REGION Network 3
   RUNG wire#powerrail
      Move(in := "EMS".Carrier[#Carrier].Zone, out1 => #Zone_Echo)
   END_RUNG
   // the same network as SCL:
   #Zone_Echo := "EMS".Carrier[#Carrier].Zone;
END_REGION

REGION Network 4
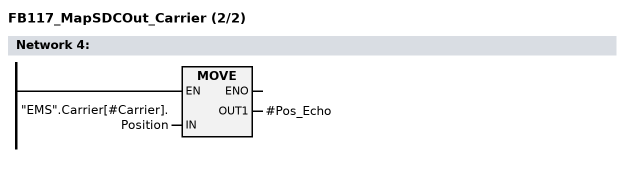
   RUNG wire#powerrail
      Move(in := "EMS".Carrier[#Carrier].Position, out1 => #Pos_Echo)
   END_RUNG
   // the same network as SCL:
   #Pos_Echo := "EMS".Carrier[#Carrier].Position;
END_REGION
END_FUNCTION_BLOCK

FUNCTION_BLOCK "FB118_TCMapSDCOut"   // FB118, LAD
{ S7_Optimized_Access := 'TRUE' }
VERSION : 0.1
   VAR_INPUT
      TC_ZoneMotion : "UDT_TC_ZoneMotion";
      Zone : Int;
      Carrier : Int;
   END_VAR
   VAR_OUTPUT
      SDCOUT_DriveFwdCmd : Bool;
      SDCOUT_DriveCmdSpeed : Word;
      SDCOUT_NextStopPos : DWord;
      SDCOUT_NextCarrierNum : Word;
      SDCOut_AtCmdPos : Bool;
   END_VAR
   VAR
      CarrierTempZone : Int;
      oneshot : Array[0..20] of Bool;
      oneshotneg : Bool;
      oneshot3 : Bool;
      resetlatch1 : Bool;
      DriveCmdSetup : Array[0..99] of Bool;
   END_VAR
   VAR_TEMP
      tempptrig : Bool;
   END_VAR
BEGIN

REGION Network 1
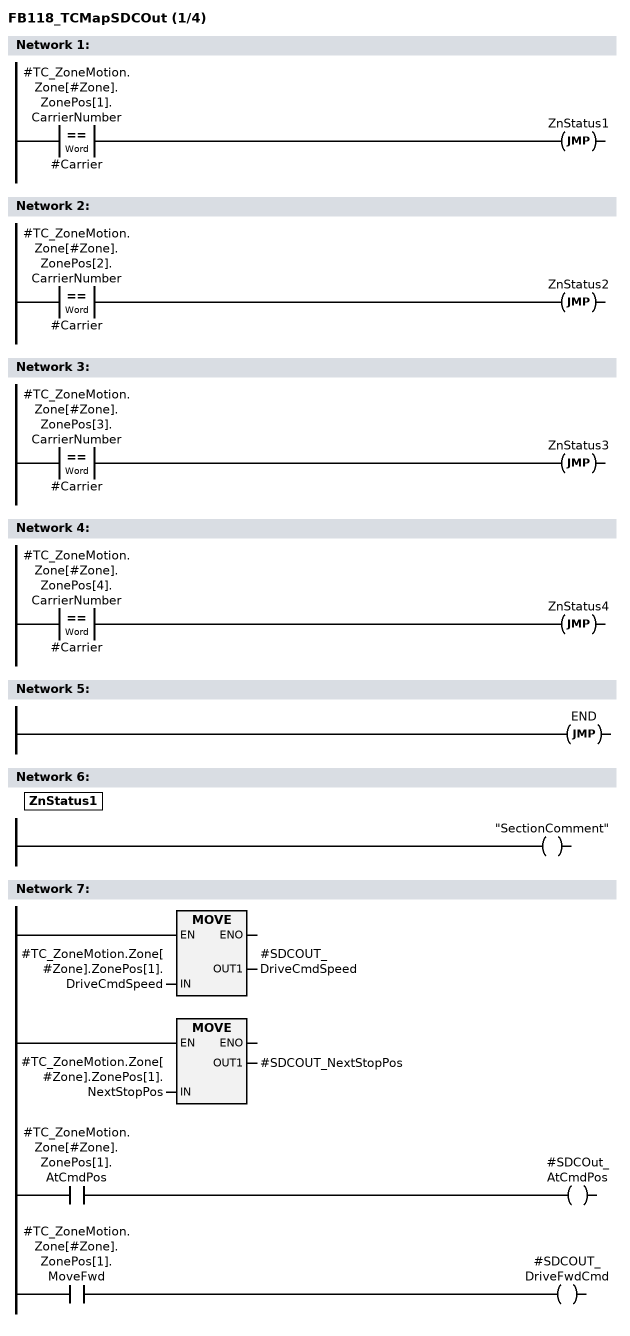
   RUNG wire#powerrail
      { S7_Templates := "SrcType := Word" } EQ_Contact(in1 := #TC_ZoneMotion.Zone[#Zone].ZonePos[1].CarrierNumber, in2 := #Carrier)
      JumpCoil( ZnStatus1 )
   END_RUNG
   // the same network as SCL:
   IF #TC_ZoneMotion.Zone[#Zone].ZonePos[1].CarrierNumber = #Carrier THEN GOTO ZnStatus1; END_IF;
END_REGION

REGION Network 2
   RUNG wire#powerrail
      { S7_Templates := "SrcType := Word" } EQ_Contact(in1 := #TC_ZoneMotion.Zone[#Zone].ZonePos[2].CarrierNumber, in2 := #Carrier)
      JumpCoil( ZnStatus2 )
   END_RUNG
   // the same network as SCL:
   IF #TC_ZoneMotion.Zone[#Zone].ZonePos[2].CarrierNumber = #Carrier THEN GOTO ZnStatus2; END_IF;
END_REGION

REGION Network 3
   RUNG wire#powerrail
      { S7_Templates := "SrcType := Word" } EQ_Contact(in1 := #TC_ZoneMotion.Zone[#Zone].ZonePos[3].CarrierNumber, in2 := #Carrier)
      JumpCoil( ZnStatus3 )
   END_RUNG
   // the same network as SCL:
   IF #TC_ZoneMotion.Zone[#Zone].ZonePos[3].CarrierNumber = #Carrier THEN GOTO ZnStatus3; END_IF;
END_REGION

REGION Network 4
   RUNG wire#powerrail
      { S7_Templates := "SrcType := Word" } EQ_Contact(in1 := #TC_ZoneMotion.Zone[#Zone].ZonePos[4].CarrierNumber, in2 := #Carrier)
      JumpCoil( ZnStatus4 )
   END_RUNG
   // the same network as SCL:
   IF #TC_ZoneMotion.Zone[#Zone].ZonePos[4].CarrierNumber = #Carrier THEN GOTO ZnStatus4; END_IF;
END_REGION

REGION Network 5
   RUNG wire#powerrail
      JumpCoil( END )
   END_RUNG
   // the same network as SCL:
   GOTO END;
END_REGION

REGION Network 6
   Label( ZnStatus1 )
   RUNG wire#powerrail
      Coil( "SectionComment" )
   END_RUNG
   // the same network as SCL:
   ZnStatus1:
   "SectionComment" := TRUE;
END_REGION

REGION Network 7
   RUNG wire#powerrail
      Move(in := #TC_ZoneMotion.Zone[#Zone].ZonePos[1].DriveCmdSpeed, out1 => #SDCOUT_DriveCmdSpeed)
   END_RUNG
   RUNG wire#powerrail
      Move(in := #TC_ZoneMotion.Zone[#Zone].ZonePos[1].NextStopPos, out1 => #SDCOUT_NextStopPos)
   END_RUNG
   RUNG wire#powerrail
      Contact( #TC_ZoneMotion.Zone[#Zone].ZonePos[1].AtCmdPos )
      Coil( #SDCOut_AtCmdPos )
   END_RUNG
   RUNG wire#powerrail
      Contact( #TC_ZoneMotion.Zone[#Zone].ZonePos[1].MoveFwd )
      Coil( #SDCOUT_DriveFwdCmd )
   END_RUNG
   // the same network as SCL:
   #SDCOUT_DriveCmdSpeed := #TC_ZoneMotion.Zone[#Zone].ZonePos[1].DriveCmdSpeed;
   #SDCOUT_NextStopPos := #TC_ZoneMotion.Zone[#Zone].ZonePos[1].NextStopPos;
   #SDCOut_AtCmdPos := #TC_ZoneMotion.Zone[#Zone].ZonePos[1].AtCmdPos;
   #SDCOUT_DriveFwdCmd := #TC_ZoneMotion.Zone[#Zone].ZonePos[1].MoveFwd;
END_REGION

REGION Network 8
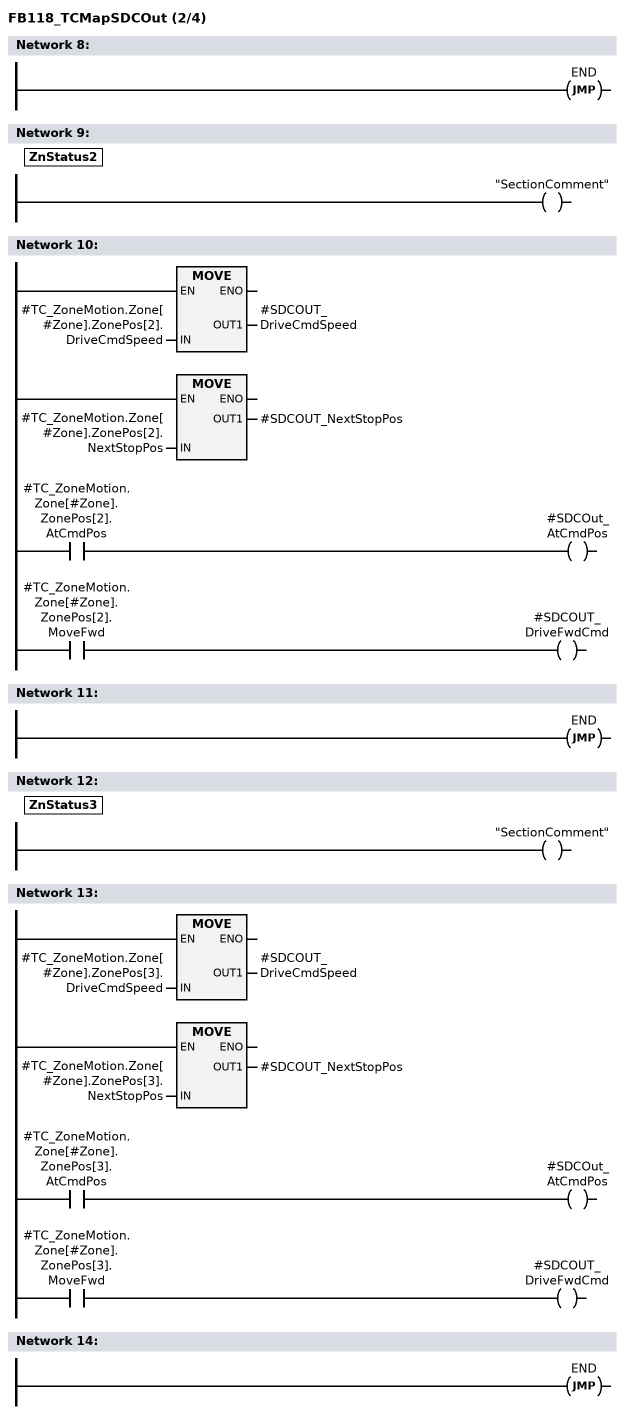
   RUNG wire#powerrail
      JumpCoil( END )
   END_RUNG
   // the same network as SCL:
   GOTO END;
END_REGION

REGION Network 9
   Label( ZnStatus2 )
   RUNG wire#powerrail
      Coil( "SectionComment" )
   END_RUNG
   // the same network as SCL:
   ZnStatus2:
   "SectionComment" := TRUE;
END_REGION

REGION Network 10
   RUNG wire#powerrail
      Move(in := #TC_ZoneMotion.Zone[#Zone].ZonePos[2].DriveCmdSpeed, out1 => #SDCOUT_DriveCmdSpeed)
   END_RUNG
   RUNG wire#powerrail
      Move(in := #TC_ZoneMotion.Zone[#Zone].ZonePos[2].NextStopPos, out1 => #SDCOUT_NextStopPos)
   END_RUNG
   RUNG wire#powerrail
      Contact( #TC_ZoneMotion.Zone[#Zone].ZonePos[2].AtCmdPos )
      Coil( #SDCOut_AtCmdPos )
   END_RUNG
   RUNG wire#powerrail
      Contact( #TC_ZoneMotion.Zone[#Zone].ZonePos[2].MoveFwd )
      Coil( #SDCOUT_DriveFwdCmd )
   END_RUNG
   // the same network as SCL:
   #SDCOUT_DriveCmdSpeed := #TC_ZoneMotion.Zone[#Zone].ZonePos[2].DriveCmdSpeed;
   #SDCOUT_NextStopPos := #TC_ZoneMotion.Zone[#Zone].ZonePos[2].NextStopPos;
   #SDCOut_AtCmdPos := #TC_ZoneMotion.Zone[#Zone].ZonePos[2].AtCmdPos;
   #SDCOUT_DriveFwdCmd := #TC_ZoneMotion.Zone[#Zone].ZonePos[2].MoveFwd;
END_REGION

REGION Network 11
   RUNG wire#powerrail
      JumpCoil( END )
   END_RUNG
   // the same network as SCL:
   GOTO END;
END_REGION

REGION Network 12
   Label( ZnStatus3 )
   RUNG wire#powerrail
      Coil( "SectionComment" )
   END_RUNG
   // the same network as SCL:
   ZnStatus3:
   "SectionComment" := TRUE;
END_REGION

REGION Network 13
   RUNG wire#powerrail
      Move(in := #TC_ZoneMotion.Zone[#Zone].ZonePos[3].DriveCmdSpeed, out1 => #SDCOUT_DriveCmdSpeed)
   END_RUNG
   RUNG wire#powerrail
      Move(in := #TC_ZoneMotion.Zone[#Zone].ZonePos[3].NextStopPos, out1 => #SDCOUT_NextStopPos)
   END_RUNG
   RUNG wire#powerrail
      Contact( #TC_ZoneMotion.Zone[#Zone].ZonePos[3].AtCmdPos )
      Coil( #SDCOut_AtCmdPos )
   END_RUNG
   RUNG wire#powerrail
      Contact( #TC_ZoneMotion.Zone[#Zone].ZonePos[3].MoveFwd )
      Coil( #SDCOUT_DriveFwdCmd )
   END_RUNG
   // the same network as SCL:
   #SDCOUT_DriveCmdSpeed := #TC_ZoneMotion.Zone[#Zone].ZonePos[3].DriveCmdSpeed;
   #SDCOUT_NextStopPos := #TC_ZoneMotion.Zone[#Zone].ZonePos[3].NextStopPos;
   #SDCOut_AtCmdPos := #TC_ZoneMotion.Zone[#Zone].ZonePos[3].AtCmdPos;
   #SDCOUT_DriveFwdCmd := #TC_ZoneMotion.Zone[#Zone].ZonePos[3].MoveFwd;
END_REGION

REGION Network 14
   RUNG wire#powerrail
      JumpCoil( END )
   END_RUNG
   // the same network as SCL:
   GOTO END;
END_REGION

REGION Network 15
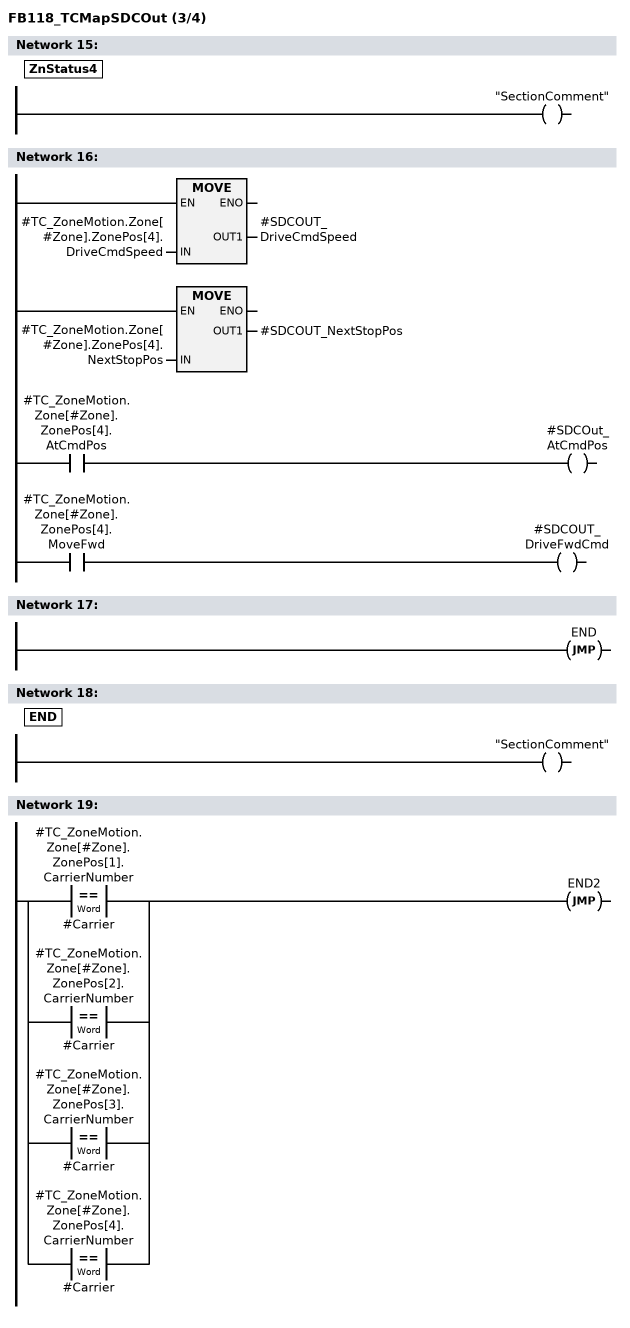
   Label( ZnStatus4 )
   RUNG wire#powerrail
      Coil( "SectionComment" )
   END_RUNG
   // the same network as SCL:
   ZnStatus4:
   "SectionComment" := TRUE;
END_REGION

REGION Network 16
   RUNG wire#powerrail
      Move(in := #TC_ZoneMotion.Zone[#Zone].ZonePos[4].DriveCmdSpeed, out1 => #SDCOUT_DriveCmdSpeed)
   END_RUNG
   RUNG wire#powerrail
      Move(in := #TC_ZoneMotion.Zone[#Zone].ZonePos[4].NextStopPos, out1 => #SDCOUT_NextStopPos)
   END_RUNG
   RUNG wire#powerrail
      Contact( #TC_ZoneMotion.Zone[#Zone].ZonePos[4].AtCmdPos )
      Coil( #SDCOut_AtCmdPos )
   END_RUNG
   RUNG wire#powerrail
      Contact( #TC_ZoneMotion.Zone[#Zone].ZonePos[4].MoveFwd )
      Coil( #SDCOUT_DriveFwdCmd )
   END_RUNG
   // the same network as SCL:
   #SDCOUT_DriveCmdSpeed := #TC_ZoneMotion.Zone[#Zone].ZonePos[4].DriveCmdSpeed;
   #SDCOUT_NextStopPos := #TC_ZoneMotion.Zone[#Zone].ZonePos[4].NextStopPos;
   #SDCOut_AtCmdPos := #TC_ZoneMotion.Zone[#Zone].ZonePos[4].AtCmdPos;
   #SDCOUT_DriveFwdCmd := #TC_ZoneMotion.Zone[#Zone].ZonePos[4].MoveFwd;
END_REGION

REGION Network 17
   RUNG wire#powerrail
      JumpCoil( END )
   END_RUNG
   // the same network as SCL:
   GOTO END;
END_REGION

REGION Network 18
   Label( END )
   RUNG wire#powerrail
      Coil( "SectionComment" )
   END_RUNG
   // the same network as SCL:
   END:
   "SectionComment" := TRUE;
END_REGION

REGION Network 19
   RUNG wire#powerrail
      { S7_Templates := "SrcType := Word" } EQ_Contact(in1 := #TC_ZoneMotion.Zone[#Zone].ZonePos[1].CarrierNumber, in2 := #Carrier)
      wire#w1
      JumpCoil( END2 )
   END_RUNG
   RUNG wire#powerrail
      { S7_Templates := "SrcType := Word" } EQ_Contact(in1 := #TC_ZoneMotion.Zone[#Zone].ZonePos[2].CarrierNumber, in2 := #Carrier)
   END_RUNG wire#w1
   RUNG wire#powerrail
      { S7_Templates := "SrcType := Word" } EQ_Contact(in1 := #TC_ZoneMotion.Zone[#Zone].ZonePos[3].CarrierNumber, in2 := #Carrier)
   END_RUNG wire#w1
   RUNG wire#powerrail
      { S7_Templates := "SrcType := Word" } EQ_Contact(in1 := #TC_ZoneMotion.Zone[#Zone].ZonePos[4].CarrierNumber, in2 := #Carrier)
   END_RUNG wire#w1
   // the same network as SCL:
   IF (#TC_ZoneMotion.Zone[#Zone].ZonePos[1].CarrierNumber = #Carrier) OR (#TC_ZoneMotion.Zone[#Zone].ZonePos[2].CarrierNumber = #Carrier) OR (#TC_ZoneMotion.Zone[#Zone].ZonePos[3].CarrierNumber = #Carrier) OR (#TC_ZoneMotion.Zone[#Zone].ZonePos[4].CarrierNumber = #Carrier) THEN
       GOTO END2;
   END_IF;
END_REGION

REGION Network 20
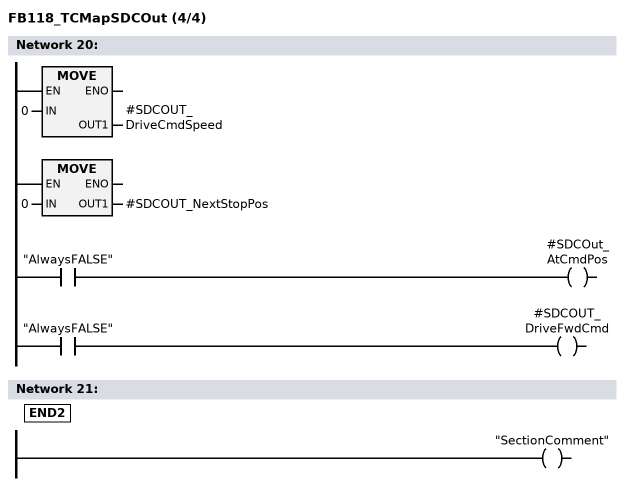
   RUNG wire#powerrail
      Move(in := 0, out1 => #SDCOUT_DriveCmdSpeed)
   END_RUNG
   RUNG wire#powerrail
      Move(in := 0, out1 => #SDCOUT_NextStopPos)
   END_RUNG
   RUNG wire#powerrail
      Contact( "AlwaysFALSE" )
      Coil( #SDCOut_AtCmdPos )
   END_RUNG
   RUNG wire#powerrail
      Contact( "AlwaysFALSE" )
      Coil( #SDCOUT_DriveFwdCmd )
   END_RUNG
   // the same network as SCL:
   #SDCOUT_DriveCmdSpeed := 0;
   #SDCOUT_NextStopPos := 0;
   #SDCOut_AtCmdPos := "AlwaysFALSE";
   #SDCOUT_DriveFwdCmd := "AlwaysFALSE";
END_REGION

REGION Network 21
   Label( END2 )
   RUNG wire#powerrail
      Coil( "SectionComment" )
   END_RUNG
   // the same network as SCL:
   END2:
   "SectionComment" := TRUE;
END_REGION
END_FUNCTION_BLOCK

FUNCTION_BLOCK "FB119_ZoneTrafficCop"   // FB119, LAD
{ S7_Optimized_Access := 'FALSE' }
VERSION : 0.1
   VAR_INPUT
      EMS : "UDT_System";
      Zone : Int := 1;
   END_VAR
   VAR_OUTPUT
      TrafficCopZone : "UDT_TrafficCopZoneStructure";
   END_VAR
   VAR
      SectionComment : Bool;
      TotalZonePositions : Int;
   END_VAR
BEGIN

REGION Network 1: Section Comment
   // Section Logic for Current Carrier number in Position 1 - Max Carrier in Zone Position Array
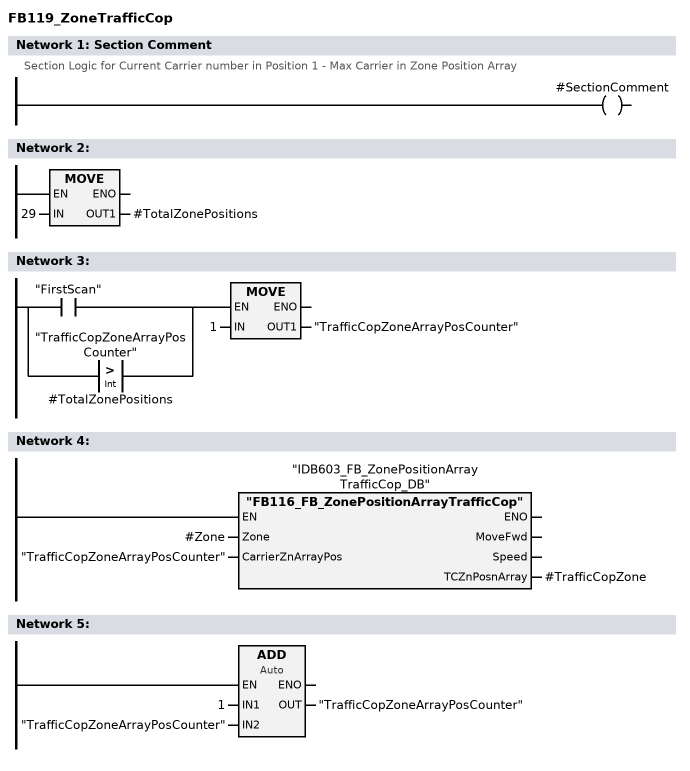
   RUNG wire#powerrail
      Coil( #SectionComment )
   END_RUNG
   // the same network as SCL:
   #SectionComment := TRUE;
END_REGION

REGION Network 2
   RUNG wire#powerrail
      Move(in := 29, out1 => #TotalZonePositions)
   END_RUNG
   // the same network as SCL:
   #TotalZonePositions := 29;
END_REGION

REGION Network 3
   RUNG wire#powerrail
      Contact( "FirstScan" )
      wire#w1
      Move(in := 1, out1 => "TrafficCopZoneArrayPosCounter")
   END_RUNG
   RUNG wire#powerrail
      { S7_Templates := "SrcType := Int" } GT_Contact(in1 := "TrafficCopZoneArrayPosCounter", in2 := #TotalZonePositions)
   END_RUNG wire#w1
   // the same network as SCL:
   IF "FirstScan" OR ("TrafficCopZoneArrayPosCounter" > #TotalZonePositions) THEN
       "TrafficCopZoneArrayPosCounter" := 1;
   END_IF;
END_REGION

REGION Network 4
   RUNG wire#powerrail
      "IDB603_FB_ZonePositionArrayTrafficCop_DB"(Zone := #Zone, CarrierZnArrayPos := "TrafficCopZoneArrayPosCounter", MoveFwd =>, Speed =>, TCZnPosnArray => #TrafficCopZone)
   END_RUNG
   // the same network as SCL:
   "IDB603_FB_ZonePositionArrayTrafficCop_DB"(Zone := #Zone,   // "FB116_FB_ZonePositionArrayTrafficCop"
                           CarrierZnArrayPos := "TrafficCopZoneArrayPosCounter",
                           TCZnPosnArray => #TrafficCopZone);
END_REGION

REGION Network 5
   RUNG wire#powerrail
      Add(in1 := 1, in2 := "TrafficCopZoneArrayPosCounter", out => "TrafficCopZoneArrayPosCounter")
   END_RUNG
   // the same network as SCL:
   "TrafficCopZoneArrayPosCounter" := 1 + "TrafficCopZoneArrayPosCounter";
END_REGION
END_FUNCTION_BLOCK

FUNCTION_BLOCK "FB120_ZoneSpacingCheck"   // FB120, SCL
{ S7_Optimized_Access := 'TRUE' }
VERSION : 0.1
   VAR_INPUT
      Zone : Int;
      TotalPosition : Int;
      EMS : "UDT_System";
   END_VAR
   VAR_OUTPUT
      GapSpacingFault : Bool;
      GapFaultZnPosition : Int;
      FirstCarrierNumGapFlt : Int;
      SecondCarrierNumGapFlt : Int;
   END_VAR
   VAR_TEMP
      ZnPosCounter : Int;
      ZoneFound : Word;
      FirstHighPos : Int;
      FirstLowPos : Int;
      NextLowPos : Int;
      NextHighPos : Int;
      GapSpaceActual : Int;
      GapSpaceActualhiLimit : Int;
      GapSpaceActualLowLimit : Int;
      NextZnPosCounter : Int;
      MaxGapSpacing : Int;
   END_VAR
BEGIN
       #ZnPosCounter := 1;
       #GapSpacingFault := 0;
       #GapFaultZnPosition := 0;
       #FirstCarrierNumGapFlt := 0;
       #SecondCarrierNumGapFlt := 0;
       FOR #ZnPosCounter := 1 TO #TotalPosition DO
           #NextZnPosCounter := #ZnPosCounter + 1;
           IF #EMS.Zone[#Zone].CarrierZnStatus[#NextZnPosCounter].CarrierNumber = 0 THEN
               ;
               RETURN;
           END_IF;

           #GapSpaceActual := #EMS.Zone[#Zone].CarrierZnStatus[#ZnPosCounter].Position - #EMS.Zone[#Zone].CarrierZnStatus[#NextZnPosCounter].Position;
           #MaxGapSpacing := #GapSpaceActual + #EMS.Zone[#Zone].InPositionTolerance;
           IF #EMS.Zone[#Zone].AccumZone = 1 & #MaxGapSpacing < #EMS.Zone[#Zone].CarrierSpacing OR #EMS.Zone[#Zone].ProductionZone = 1 & #MaxGapSpacing < #EMS.Zone[#Zone].ProductionZoneSpacing THEN
               #GapSpacingFault := 1;
               #GapFaultZnPosition := #ZnPosCounter;
               #FirstCarrierNumGapFlt := #EMS.Zone[#Zone].CarrierZnStatus[#ZnPosCounter].CarrierNumber;
               #SecondCarrierNumGapFlt := #EMS.Zone[#Zone].CarrierZnStatus[#NextZnPosCounter].CarrierNumber;
          ELSE
    #GapSpacingFault := 0;
     //#FirstCarrierNumGapFlt := 0;
     //#SecondCarrierNumGapFlt := 0;
               RETURN;
           END_IF;
       END_FOR;
END_FUNCTION_BLOCK

// folder: 04_FCs

FUNCTION "FC100_EMS_System" : Void   // FC100, LAD
{ S7_Optimized_Access := 'TRUE' }
VERSION : 0.1
   VAR_TEMP
      TEMPCARRIERNUMBR : Word;
   END_VAR
BEGIN

REGION Network 1
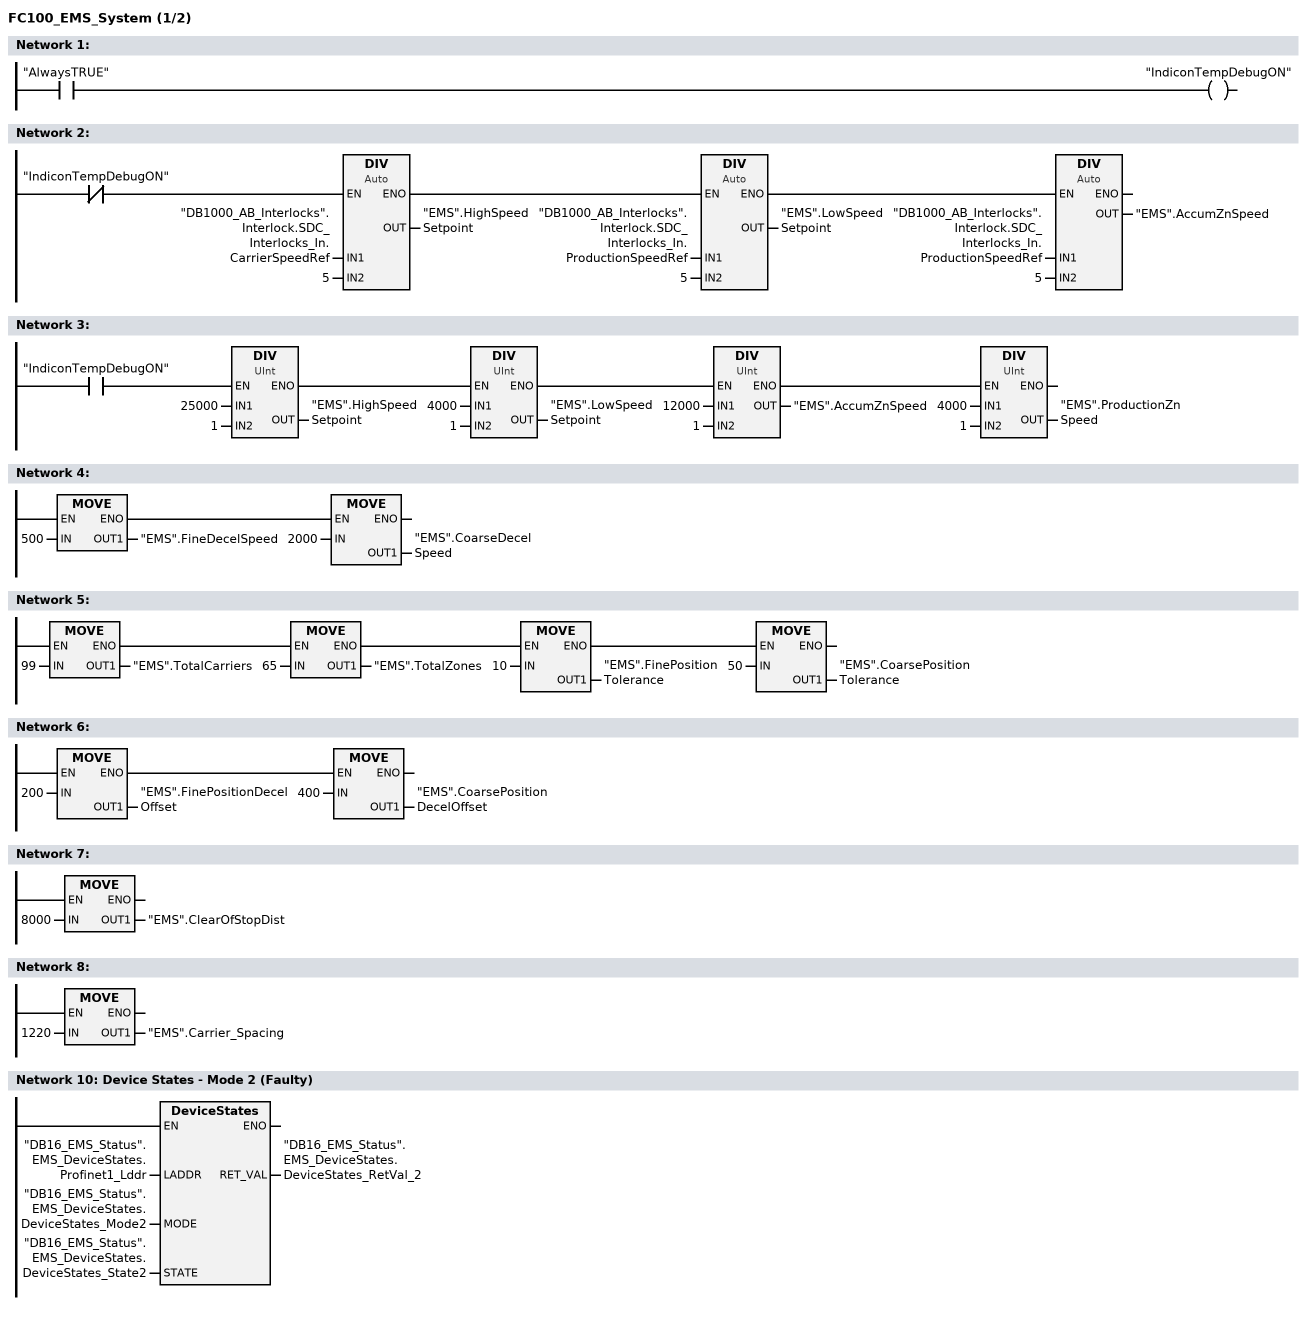
   RUNG wire#powerrail
      Contact( "AlwaysTRUE" )
      Coil( "IndiconTempDebugON" )
   END_RUNG
   // the same network as SCL:
   "IndiconTempDebugON" := "AlwaysTRUE";
END_REGION

REGION Network 2
   RUNG wire#powerrail
      I_Contact( "IndiconTempDebugON" )
      Div(in1 := "DB1000_AB_Interlocks".Interlock.SDC_Interlocks_In.CarrierSpeedRef, in2 := 5, out => "EMS".HighSpeedSetpoint)
      Div(in1 := "DB1000_AB_Interlocks".Interlock.SDC_Interlocks_In.ProductionSpeedRef, in2 := 5, out => "EMS".LowSpeedSetpoint)
      Div(in1 := "DB1000_AB_Interlocks".Interlock.SDC_Interlocks_In.ProductionSpeedRef, in2 := 5, out => "EMS".AccumZnSpeed)
   END_RUNG
   // the same network as SCL:
   IF NOT "IndiconTempDebugON" THEN
       "EMS".HighSpeedSetpoint := "DB1000_AB_Interlocks".Interlock.SDC_Interlocks_In.CarrierSpeedRef / 5;
       "EMS".LowSpeedSetpoint := "DB1000_AB_Interlocks".Interlock.SDC_Interlocks_In.ProductionSpeedRef / 5;
       "EMS".AccumZnSpeed := "DB1000_AB_Interlocks".Interlock.SDC_Interlocks_In.ProductionSpeedRef / 5;
   END_IF;
END_REGION

REGION Network 3
   RUNG wire#powerrail
      Contact( "IndiconTempDebugON" )
      { S7_Templates := "SrcType := UInt" } Div(in1 := 25000, in2 := 1, out => "EMS".HighSpeedSetpoint)
      { S7_Templates := "SrcType := UInt" } Div(in1 := 4000, in2 := 1, out => "EMS".LowSpeedSetpoint)
      { S7_Templates := "SrcType := UInt" } Div(in1 := 12000, in2 := 1, out => "EMS".AccumZnSpeed)
      { S7_Templates := "SrcType := UInt" } Div(in1 := 4000, in2 := 1, out => "EMS".ProductionZnSpeed)
   END_RUNG
   // the same network as SCL:
   IF "IndiconTempDebugON" THEN
       "EMS".HighSpeedSetpoint := 25000 / 1;
       "EMS".LowSpeedSetpoint := 4000 / 1;
       "EMS".AccumZnSpeed := 12000 / 1;
       "EMS".ProductionZnSpeed := 4000 / 1;
   END_IF;
END_REGION

REGION Network 4
   RUNG wire#powerrail
      Move(in := 500, out1 => "EMS".FineDecelSpeed)
      Move(in := 2000, out1 => "EMS".CoarseDecelSpeed)
   END_RUNG
   // the same network as SCL:
   "EMS".FineDecelSpeed := 500;
   "EMS".CoarseDecelSpeed := 2000;
END_REGION

REGION Network 5
   RUNG wire#powerrail
      Move(in := 99, out1 => "EMS".TotalCarriers)
      Move(in := 65, out1 => "EMS".TotalZones)
      Move(in := 10, out1 => "EMS".FinePositionTolerance)
      Move(in := 50, out1 => "EMS".CoarsePositionTolerance)
   END_RUNG
   // the same network as SCL:
   "EMS".TotalCarriers := 99;
   "EMS".TotalZones := 65;
   "EMS".FinePositionTolerance := 10;
   "EMS".CoarsePositionTolerance := 50;
END_REGION

REGION Network 6
   RUNG wire#powerrail
      Move(in := 200, out1 => "EMS".FinePositionDecelOffset)
      Move(in := 400, out1 => "EMS".CoarsePositionDecelOffset)
   END_RUNG
   // the same network as SCL:
   "EMS".FinePositionDecelOffset := 200;
   "EMS".CoarsePositionDecelOffset := 400;
END_REGION

REGION Network 7
   RUNG wire#powerrail
      Move(in := 8000, out1 => "EMS".ClearOfStopDist)
   END_RUNG
   // the same network as SCL:
   "EMS".ClearOfStopDist := 8000;
END_REGION

REGION Network 8
   RUNG wire#powerrail
      Move(in := 1220, out1 => "EMS".Carrier_Spacing)
   END_RUNG
   // the same network as SCL:
   "EMS".Carrier_Spacing := 1220;
END_REGION

REGION Network 10: Device States - Mode 2 (Faulty)
   // no SCL statement known for DeviceStates: written as a call
   "DB16_EMS_Status".EMS_DeviceStates.DeviceStates_RetVal_2 := DeviceStates(LADDR := "DB16_EMS_Status".EMS_DeviceStates.Profinet1_Lddr,
                           MODE := "DB16_EMS_Status".EMS_DeviceStates.DeviceStates_Mode2,
                           STATE := "DB16_EMS_Status".EMS_DeviceStates.DeviceStates_State2);
END_REGION

REGION Network 11: Device States - Mode 4 (Exists)
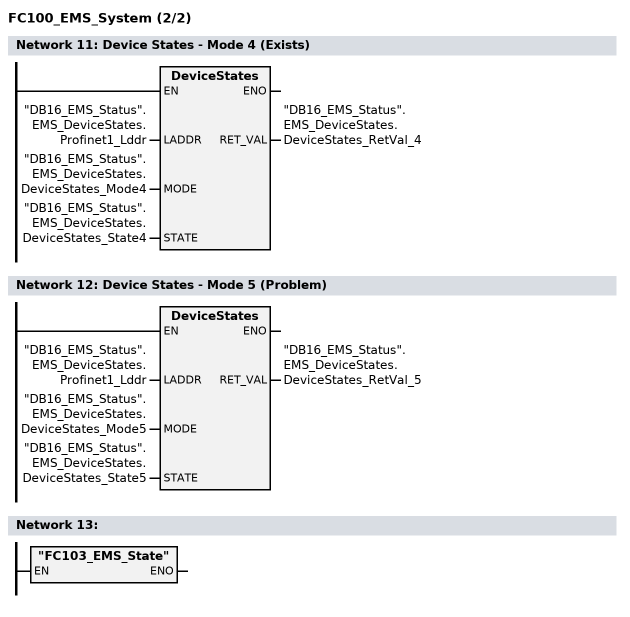
   // no SCL statement known for DeviceStates: written as a call
   "DB16_EMS_Status".EMS_DeviceStates.DeviceStates_RetVal_4 := DeviceStates(LADDR := "DB16_EMS_Status".EMS_DeviceStates.Profinet1_Lddr,
                           MODE := "DB16_EMS_Status".EMS_DeviceStates.DeviceStates_Mode4,
                           STATE := "DB16_EMS_Status".EMS_DeviceStates.DeviceStates_State4);
END_REGION

REGION Network 12: Device States - Mode 5 (Problem)
   // no SCL statement known for DeviceStates: written as a call
   "DB16_EMS_Status".EMS_DeviceStates.DeviceStates_RetVal_5 := DeviceStates(LADDR := "DB16_EMS_Status".EMS_DeviceStates.Profinet1_Lddr,
                           MODE := "DB16_EMS_Status".EMS_DeviceStates.DeviceStates_Mode5,
                           STATE := "DB16_EMS_Status".EMS_DeviceStates.DeviceStates_State5);
END_REGION

REGION Network 13
   RUNG wire#powerrail
      "FC103_EMS_State"()
   END_RUNG
   // the same network as SCL:
   "FC103_EMS_State"();
END_REGION
END_FUNCTION

FUNCTION "FC101_SystemZoneFind" : Void   // FC101, LAD
{ S7_Optimized_Access := 'FALSE' }
VERSION : 0.1
   VAR_TEMP
      resettemp : Bool;
      dntemp : Bool;
   END_VAR
BEGIN

REGION Network 1
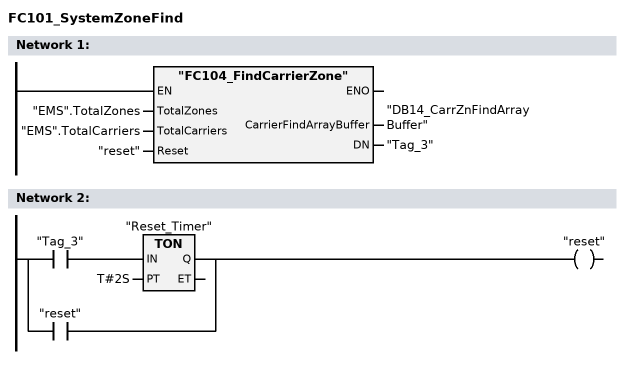
   RUNG wire#powerrail
      "FC104_FindCarrierZone"(TotalZones := "EMS".TotalZones, TotalCarriers := "EMS".TotalCarriers, Reset := "reset", CarrierFindArrayBuffer => "DB14_CarrZnFindArrayBuffer", DN => "Tag_3")
   END_RUNG
   // the same network as SCL:
   "FC104_FindCarrierZone"(TotalZones := "EMS".TotalZones,
                           TotalCarriers := "EMS".TotalCarriers,
                           Reset := "reset",
                           CarrierFindArrayBuffer => "DB14_CarrZnFindArrayBuffer",
                           DN => "Tag_3");
END_REGION

REGION Network 2
   "Reset_Timer".TON(IN := "Tag_3", PT := T#2S);
   "reset" := "Reset_Timer".Q OR "reset";
END_REGION
END_FUNCTION

FUNCTION "FC102_CarrierSetup" : Void   // FC102, LAD
{ S7_Optimized_Access := 'FALSE' }
VERSION : 0.1
   VAR_TEMP
      CarrierCounter : Int;
      TotalCarriers : Int;
      CounterReset : Bool;
      CarrierCounterDN : Bool;
      OneShotClock_2hz : Bool;
   END_VAR
BEGIN

REGION Network 1
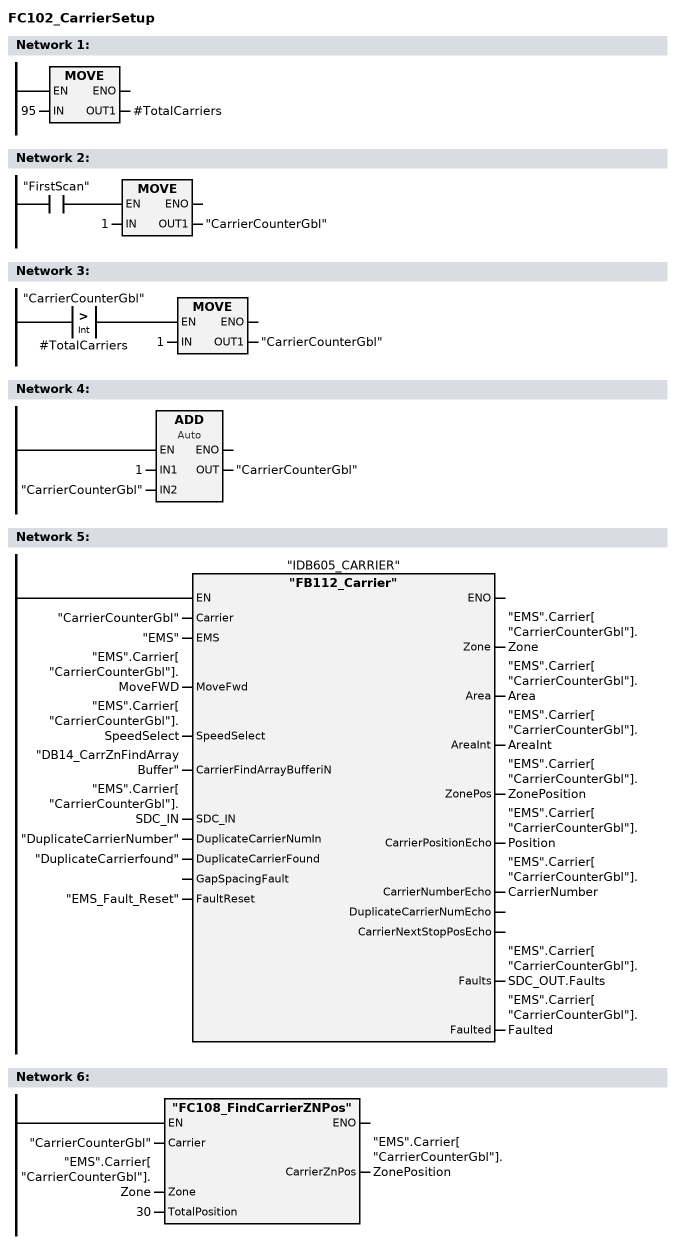
   RUNG wire#powerrail
      Move(in := 95, out1 => #TotalCarriers)
   END_RUNG
   // the same network as SCL:
   #TotalCarriers := 95;
END_REGION

REGION Network 2
   RUNG wire#powerrail
      Contact( "FirstScan" )
      Move(in := 1, out1 => "CarrierCounterGbl")
   END_RUNG
   // the same network as SCL:
   IF "FirstScan" THEN "CarrierCounterGbl" := 1; END_IF;
END_REGION

REGION Network 3
   RUNG wire#powerrail
      { S7_Templates := "SrcType := Int" } GT_Contact(in1 := "CarrierCounterGbl", in2 := #TotalCarriers)
      Move(in := 1, out1 => "CarrierCounterGbl")
   END_RUNG
   // the same network as SCL:
   IF "CarrierCounterGbl" > #TotalCarriers THEN "CarrierCounterGbl" := 1; END_IF;
END_REGION

REGION Network 4
   RUNG wire#powerrail
      Add(in1 := 1, in2 := "CarrierCounterGbl", out => "CarrierCounterGbl")
   END_RUNG
   // the same network as SCL:
   "CarrierCounterGbl" := 1 + "CarrierCounterGbl";
END_REGION

REGION Network 5
   RUNG wire#powerrail
      "IDB605_CARRIER"(Carrier := "CarrierCounterGbl", EMS := "EMS", MoveFwd := "EMS".Carrier["CarrierCounterGbl"].MoveFWD, SpeedSelect := "EMS".Carrier["CarrierCounterGbl"].SpeedSelect, CarrierFindArrayBufferiN := "DB14_CarrZnFindArrayBuffer", SDC_IN := "EMS".Carrier["CarrierCounterGbl"].SDC_IN, DuplicateCarrierNumIn := "DuplicateCarrierNumber", DuplicateCarrierFound := "DuplicateCarrierfound", GapSpacingFault :=, FaultReset := "EMS_Fault_Reset", Zone => "EMS".Carrier["CarrierCounterGbl"].Zone, Area => "EMS".Carrier["CarrierCounterGbl"].Area, AreaInt => "EMS".Carrier["CarrierCounterGbl"].AreaInt, ZonePos => "EMS".Carrier["CarrierCounterGbl"].ZonePosition, CarrierPositionEcho => "EMS".Carrier["CarrierCounterGbl"].Position, CarrierNumberEcho => "EMS".Carrier["CarrierCounterGbl"].CarrierNumber, DuplicateCarrierNumEcho =>, CarrierNextStopPosEcho =>, Faults => "EMS".Carrier["CarrierCounterGbl"].SDC_OUT.Faults, Faulted => "EMS".Carrier["CarrierCounterGbl"].Faulted)
   END_RUNG
   // the same network as SCL:
   "IDB605_CARRIER"(Carrier := "CarrierCounterGbl",   // "FB112_Carrier"
                    EMS := "EMS",
                    MoveFwd := "EMS".Carrier["CarrierCounterGbl"].MoveFWD,
                    SpeedSelect := "EMS".Carrier["CarrierCounterGbl"].SpeedSelect,
                    CarrierFindArrayBufferiN := "DB14_CarrZnFindArrayBuffer",
                    SDC_IN := "EMS".Carrier["CarrierCounterGbl"].SDC_IN,
                    DuplicateCarrierNumIn := "DuplicateCarrierNumber",
                    DuplicateCarrierFound := "DuplicateCarrierfound",
                    FaultReset := "EMS_Fault_Reset",
                    Zone => "EMS".Carrier["CarrierCounterGbl"].Zone,
                    Area => "EMS".Carrier["CarrierCounterGbl"].Area,
                    AreaInt => "EMS".Carrier["CarrierCounterGbl"].AreaInt,
                    ZonePos => "EMS".Carrier["CarrierCounterGbl"].ZonePosition,
                    CarrierPositionEcho => "EMS".Carrier["CarrierCounterGbl"].Position,
                    CarrierNumberEcho => "EMS".Carrier["CarrierCounterGbl"].CarrierNumber,
                    Faults => "EMS".Carrier["CarrierCounterGbl"].SDC_OUT.Faults,
                    Faulted => "EMS".Carrier["CarrierCounterGbl"].Faulted);
END_REGION

REGION Network 6
   RUNG wire#powerrail
      "FC108_FindCarrierZNPos"(Carrier := "CarrierCounterGbl", Zone := "EMS".Carrier["CarrierCounterGbl"].Zone, TotalPosition := 30, CarrierZnPos => "EMS".Carrier["CarrierCounterGbl"].ZonePosition)
   END_RUNG
   // the same network as SCL:
   "FC108_FindCarrierZNPos"(Carrier := "CarrierCounterGbl",
                           Zone := "EMS".Carrier["CarrierCounterGbl"].Zone,
                           TotalPosition := 30,
                           CarrierZnPos => "EMS".Carrier["CarrierCounterGbl"].ZonePosition);
END_REGION
END_FUNCTION

FUNCTION "FC103_EMS_State" : Void   // FC103, SCL
{ S7_Optimized_Access := 'TRUE' }
VERSION : 0.1
   VAR_TEMP
      N : Int;
   END_VAR
BEGIN
   FOR #N := 1 TO 82 DO
       // Statement section FOR
       IF "DB16_EMS_Status".EMS_DeviceStates.DeviceStates_State4[#N] = FALSE
       THEN
           "DB16_EMS_Status".EMS_DeviceStates.DeviceStates_Condition_HMI[#N] := 0;
       ELSE
           IF "DB16_EMS_Status".EMS_DeviceStates.DeviceStates_State4[#N] = TRUE
           THEN
               "DB16_EMS_Status".EMS_DeviceStates.DeviceStates_Condition_HMI[#N] := 1;
           END_IF;
           IF "DB16_EMS_Status".EMS_DeviceStates.DeviceStates_State5[#N] = TRUE
           THEN
               "DB16_EMS_Status".EMS_DeviceStates.DeviceStates_Condition_HMI[#N] := 3;
           END_IF;
           IF "DB16_EMS_Status".EMS_DeviceStates.DeviceStates_State2[#N] = TRUE
           THEN
               "DB16_EMS_Status".EMS_DeviceStates.DeviceStates_Condition_HMI[#N] := 2;
           END_IF;
       END_IF;

   END_FOR;
END_FUNCTION

FUNCTION "FC104_FindCarrierZone" : Void   // FC104, SCL
{ S7_Optimized_Access := 'FALSE' }
VERSION : 0.1
   VAR_INPUT
      TotalZones : Int;
      TotalCarriers : Int;
      Reset : Bool;
   END_VAR
   VAR_OUTPUT
      CarrierFindArrayBuffer : "UDT_Carrier";
      DN : Bool;
   END_VAR
   VAR_TEMP
      ZoneCounter : Int;
      ZoneFound : Word;
      CarrierCounter : Int;
      ZouneFound : Int;
   END_VAR
BEGIN
   //[***********************************************************************************NO EDITS*******************************************************************************************************]
   //FC200 - Find Carrier Zone
   //Double loop counter finds which zone carrier is located based on Zone Start Position and End Position and records the result in the system EMS DB for each carrier
   //- EMS.Carrier[x].Zone
   //***************************************************************************************************************************************************************************************************

      #ZoneCounter := 1;
      #CarrierCounter := 1;


       FOR #ZoneCounter := 1 TO #TotalZones DO
           // Statement section FOR
           ;
           WHILE #CarrierCounter <= #TotalCarriers DO
               ;
               IF "EMS".Carrier[#CarrierCounter].Position > "EMS".Zone[#ZoneCounter].StartPos AND
                   "EMS".Carrier[#CarrierCounter].Position < "EMS".Zone[#ZoneCounter].EndPos
               THEN
                   #CarrierFindArrayBuffer.CARRIER[#CarrierCounter].Zone := #ZoneCounter;
                   #CarrierFindArrayBuffer.CARRIER[#CarrierCounter].Area := "EMS".Zone[#ZoneCounter].Area;

               END_IF;

               #CarrierCounter := #CarrierCounter + 1;
               "cARIERLOOPCOUNT2" := #CarrierCounter;
           END_WHILE;
           #CarrierCounter := 1;
           "ZoneCnt" := #ZoneCounter;
       END_FOR;
END_FUNCTION

FUNCTION "FC105_ZoneCarrierStatus" : Void   // FC105, SCL
{ S7_Optimized_Access := 'FALSE' }
VERSION : 0.1
   VAR_INPUT
      Zone : Int;
      TotalPosition : Int;
      TotalCarriers : Int;
      TotalZones : Int;
      Reset : Bool;
   END_VAR
   VAR_OUTPUT
      ZonePosnArrayBuffer : Array[0..60] of "UDT_ZoneCarrierStatus";
      DN : Bool;
   END_VAR
   VAR_TEMP
      ZoneCounter : Int;
      ZoneFound : Word;
      CarrierCounter : Int;
      SortArrayIndex : Int;
      ArrayIndex : Int;
      Idx1 : Int;
      MaxVal : Int;
      MaxIdx1 : Int;
      Max : Int;
      Idx2 : Int;
      SelectionSort : Int;
   END_VAR
BEGIN
       //[***********************************************************************************NO EDITS*******************************************************************************************************]
       //FC201 - Find Carrier Status
       //Double loop counter finds which zone carrier is located based on Zone Start Position and End Position and records the result in the system EMS DB for each carrier
       //- EMS.Carrier[x].Zone
       //***************************************************************************************************************************************************************************************************

       #CarrierCounter := 1;
       #ArrayIndex := 1;

           WHILE #CarrierCounter <= #TotalCarriers DO
               IF "EMS".Carrier[#CarrierCounter].Zone = #Zone THEN
                   #ZonePosnArrayBuffer[#ArrayIndex].CarrierNumber := "EMS".Carrier[#CarrierCounter].SDC_IN.CarrierNumber;
                   #ZonePosnArrayBuffer[#ArrayIndex].Position := "EMS".Carrier[#CarrierCounter].Position;
                    #ArrayIndex := #ArrayIndex + 1;
                    "IndexArraytemp" := #ArrayIndex;
               ELSE
                   #ZonePosnArrayBuffer[#ArrayIndex].CarrierNumber := 0;
                   #ZonePosnArrayBuffer[#ArrayIndex].Position := 0;
               END_IF;
               #CarrierCounter := #CarrierCounter + 1;
           END_WHILE;
END_FUNCTION

FUNCTION "FC106_ZoneCarrierSort" : Void   // FC106, SCL
{ S7_Optimized_Access := 'FALSE' }
VERSION : 0.1
   VAR_INPUT
      ArrayInUnsort : Array[0..60] of "UDT_ZoneCarrierStatus";
      Max : Int;
   END_VAR
   VAR_OUTPUT
      ZonePositionArrayOut : Array[0..60] of "UDT_ZoneCarrierStatus";
   END_VAR
   VAR_TEMP
      Idx1 : Int;
      MaxVal : DWord;
      MaxIdx1 : Int;
      Idx2 : Int;
      SelectionSort : Int;
      ArrayTemp : Array[0..60] of "UDT_ZoneCarrierStatus";
      MaxCarr : Int;
   END_VAR
BEGIN
   //[***********************************************************************************NO EDITS*******************************************************************************************************]
   //FC202 - Zone Carrier Sort
   //Double loop counter Sorts Carriers in Called Zone to place in correct sequence within  zone. Zones are divided into position based on MaxCarriers allowed in zone as set in the
   //zone setup function block.  Sorted array is used in Traffic cop zone motion control
   //- EMS.Carrier[x].Zone
   //***************************************************************************************************************************************************************************************************
   #ArrayTemp := #ArrayInUnsort;


   FOR #Idx1 := 1 TO #Max BY 1 DO

       #MaxVal := #ArrayTemp[#Idx1].Position;
       IF #ArrayTemp[#Idx1].Position = 0 THEN
           EXIT;
       ELSE
           #MaxIdx1 := #Idx1;
       END_IF;